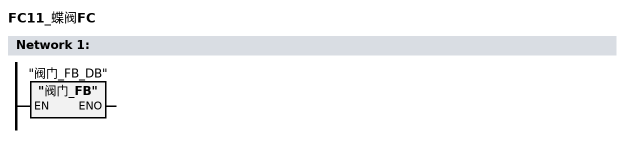
   RUNG wire#powerrail
      "阀门_FB_DB"()
   END_RUNG
   // the same network as SCL:
   "阀门_FB_DB"();   // "阀门_FB"
END_REGION
END_FUNCTION

FUNCTION "FC12_引水阀和排气阀FC" : Void   // FC12, LAD
{ S7_Optimized_Access := 'TRUE' }
VERSION : 0.1
BEGIN

REGION Network 1
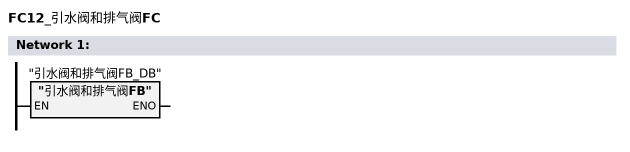
   RUNG wire#powerrail
      "引水阀和排气阀FB_DB"()
   END_RUNG
   // the same network as SCL:
   "引水阀和排气阀FB_DB"();   // "引水阀和排气阀FB"
END_REGION
END_FUNCTION

FUNCTION "FC13_电机_泵FC" : Void   // FC13, LAD
{ S7_Optimized_Access := 'TRUE' }
VERSION : 0.1
BEGIN

REGION Network 1
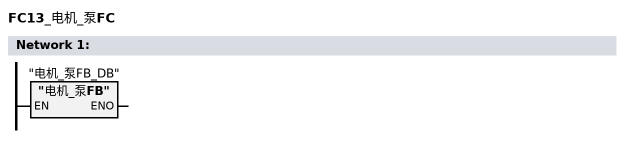
   RUNG wire#powerrail
      "电机_泵FB_DB"()
   END_RUNG
   // the same network as SCL:
   "电机_泵FB_DB"();   // "电机_泵FB"
END_REGION
END_FUNCTION

FUNCTION "FC14_DATA_ALARM" : Void   // FC14, LAD
{ S7_Optimized_Access := 'TRUE' }
VERSION : 0.1
BEGIN

REGION Network 1
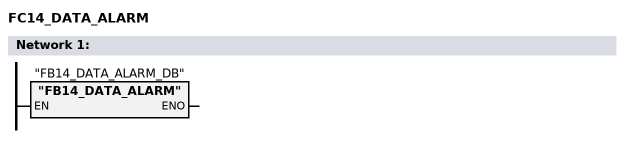
   RUNG wire#powerrail
      "FB14_DATA_ALARM_DB"()
   END_RUNG
   // the same network as SCL:
   "FB14_DATA_ALARM_DB"();   // "FB14_DATA_ALARM"
END_REGION
END_FUNCTION

FUNCTION "FC15_MOTOR_AUTO_ST" : Void   // FC15, LAD
{ S7_Optimized_Access := 'TRUE' }
VERSION : 0.1
BEGIN

REGION Network 1
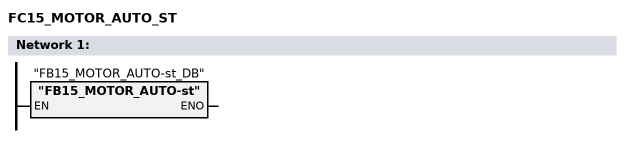
   RUNG wire#powerrail
      "FB15_MOTOR_AUTO-st_DB"()
   END_RUNG
   // the same network as SCL:
   "FB15_MOTOR_AUTO-st_DB"();   // "FB15_MOTOR_AUTO-st"
END_REGION
END_FUNCTION

FUNCTION "FC16" : Void   // FC16, LAD
{ S7_Optimized_Access := 'TRUE' }
VERSION : 0.1
   VAR_TEMP   // added for the SCL form of the ladder/FBD networks
      _w1 : Bool;
   END_VAR
BEGIN

REGION Network 1
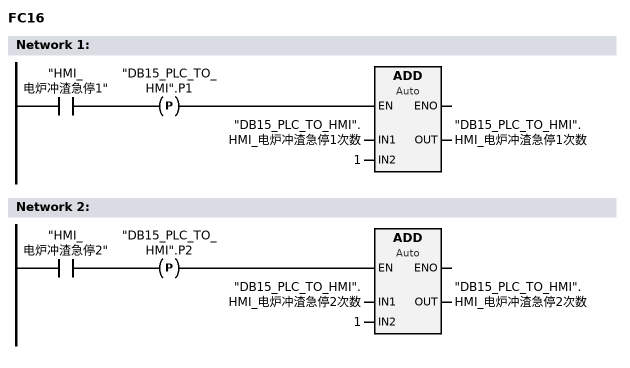
   RUNG wire#powerrail
      Contact( "HMI_电炉冲渣急停1" )
      P_Trig( "DB15_PLC_TO_HMI".P1 )
      Add(in1 := "DB15_PLC_TO_HMI".HMI_电炉冲渣急停1次数, in2 := 1, out => "DB15_PLC_TO_HMI".HMI_电炉冲渣急停1次数)
   END_RUNG
   // the same network as SCL:
   #_w1 := "HMI_电炉冲渣急停1" AND NOT "DB15_PLC_TO_HMI".P1;   // rising edge
   "DB15_PLC_TO_HMI".P1 := "HMI_电炉冲渣急停1";
   IF #_w1 THEN "DB15_PLC_TO_HMI".HMI_电炉冲渣急停1次数 := "DB15_PLC_TO_HMI".HMI_电炉冲渣急停1次数 + 1; END_IF;
END_REGION

REGION Network 2
   RUNG wire#powerrail
      Contact( "HMI_电炉冲渣急停2" )
      P_Trig( "DB15_PLC_TO_HMI".P2 )
      Add(in1 := "DB15_PLC_TO_HMI".HMI_电炉冲渣急停2次数, in2 := 1, out => "DB15_PLC_TO_HMI".HMI_电炉冲渣急停2次数)
   END_RUNG
   // the same network as SCL:
   #_w1 := "HMI_电炉冲渣急停2" AND NOT "DB15_PLC_TO_HMI".P2;   // rising edge
   "DB15_PLC_TO_HMI".P2 := "HMI_电炉冲渣急停2";
   IF #_w1 THEN "DB15_PLC_TO_HMI".HMI_电炉冲渣急停2次数 := "DB15_PLC_TO_HMI".HMI_电炉冲渣急停2次数 + 1; END_IF;
END_REGION
END_FUNCTION

ORGANIZATION_BLOCK "Main"   // OB1, LAD, ProgramCycle
TITLE = "Main Program Sweep (Cycle)"
{ S7_Optimized_Access := 'TRUE' }
VERSION : 0.1
   VAR_INPUT
      Initial_Call : Bool;   // Initial call of this OB
      Remanence : Bool;   // =True, if remanent data are available
   END_VAR
BEGIN

REGION Network 1
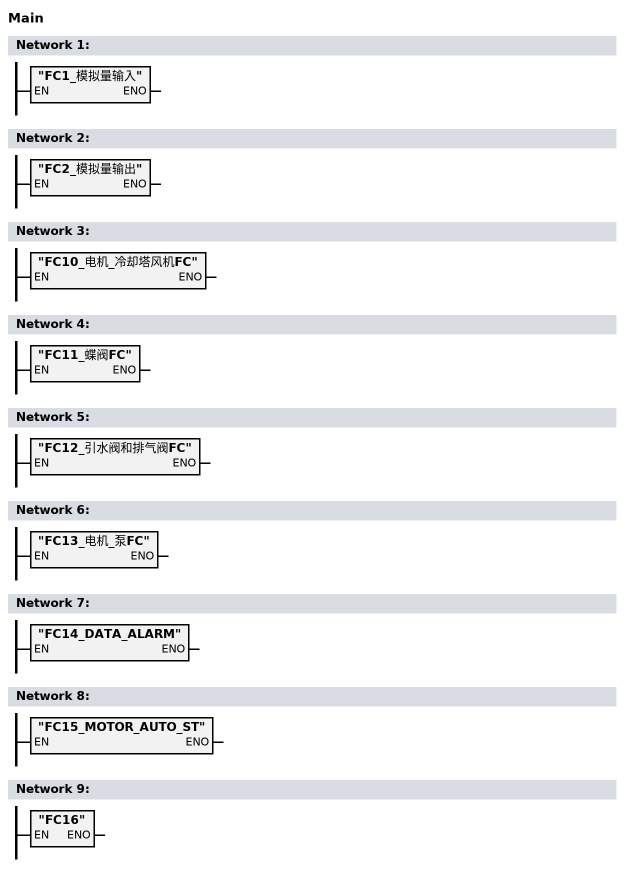
   RUNG wire#powerrail
      "FC1_模拟量输入"()
   END_RUNG
   // the same network as SCL:
   "FC1_模拟量输入"();
END_REGION

REGION Network 2
   RUNG wire#powerrail
      "FC2_模拟量输出"()
   END_RUNG
   // the same network as SCL:
   "FC2_模拟量输出"();
END_REGION

REGION Network 3
   RUNG wire#powerrail
      "FC10_电机_冷却塔风机FC"()
   END_RUNG
   // the same network as SCL:
   "FC10_电机_冷却塔风机FC"();
END_REGION

REGION Network 4
   RUNG wire#powerrail
      "FC11_蝶阀FC"()
   END_RUNG
   // the same network as SCL:
   "FC11_蝶阀FC"();
END_REGION

REGION Network 5
   RUNG wire#powerrail
      "FC12_引水阀和排气阀FC"()
   END_RUNG
   // the same network as SCL:
   "FC12_引水阀和排气阀FC"();
END_REGION

REGION Network 6
   RUNG wire#powerrail
      "FC13_电机_泵FC"()
   END_RUNG
   // the same network as SCL:
   "FC13_电机_泵FC"();
END_REGION

REGION Network 7
   RUNG wire#powerrail
      "FC14_DATA_ALARM"()
   END_RUNG
   // the same network as SCL:
   "FC14_DATA_ALARM"();
END_REGION

REGION Network 8
   RUNG wire#powerrail
      "FC15_MOTOR_AUTO_ST"()
   END_RUNG
   // the same network as SCL:
   "FC15_MOTOR_AUTO_ST"();
END_REGION

REGION Network 9
   RUNG wire#powerrail
      "FC16"()
   END_RUNG
   // the same network as SCL:
   "FC16"();
END_REGION
END_ORGANIZATION_BLOCK

ORGANIZATION_BLOCK "Cyclic interrupt"   // OB30, LAD, CyclicInterrupt
{ S7_Optimized_Access := 'TRUE' }
VERSION : 0.1
   VAR_INPUT
      Initial_Call : Bool;   // Initial call of this OB
      Event_Count : Int;   // Events discarded
   END_VAR
BEGIN
END_ORGANIZATION_BLOCK

// ===== PLC "2#SBF"  CPU 1511-1 PN =====

VAR_GLOBAL   // PLC tag table "默认变量表"
   "System_Byte" AT %MB1 : Byte;
   "FirstScan" AT %M1.0 : Bool;
   "DiagStatusUpdate" AT %M1.1 : Bool;
   "AlwaysTRUE" AT %M1.2 : Bool;
   "AlwaysFALSE" AT %M1.3 : Bool;
   "Clock_Byte" AT %MB0 : Byte;
   "Clock_10Hz" AT %M0.0 : Bool;
   "Clock_5Hz" AT %M0.1 : Bool;
   "Clock_2.5Hz" AT %M0.2 : Bool;
   "Clock_2Hz" AT %M0.3 : Bool;
   "Clock_1.25Hz" AT %M0.4 : Bool;
   "Clock_1Hz" AT %M0.5 : Bool;
   "Clock_0.625Hz" AT %M0.6 : Bool;
   "Clock_0.5Hz" AT %M0.7 : Bool;
   "1#冲渣泵本地/远程" AT %I0.0 : Bool;
   "1#冲渣泵备妥" AT %I0.1 : Bool;
   "1#冲渣泵运行" AT %I0.2 : Bool;
   "1#冲渣泵故障" AT %I0.3 : Bool;
   "2#冲渣泵本地/远程" AT %I0.4 : Bool;
   "2#冲渣泵备妥" AT %I0.5 : Bool;
   "2#冲渣泵运行" AT %I0.6 : Bool;
   "2#冲渣泵故障" AT %I0.7 : Bool;
   "3#冲渣泵本地/远程" AT %I1.0 : Bool;
   "3#冲渣泵备妥" AT %I1.1 : Bool;
   "3#冲渣泵运行" AT %I1.2 : Bool;
   "3#冲渣泵故障" AT %I1.3 : Bool;
   "4#冲渣泵本地/远程" AT %I1.4 : Bool;
   "4#冲渣泵备妥" AT %I1.5 : Bool;
   "4#冲渣泵运行" AT %I1.6 : Bool;
   "4#冲渣泵故障" AT %I1.7 : Bool;
   "5#冲渣泵本地/远程" AT %I2.0 : Bool;
   "5#冲渣泵备妥" AT %I2.1 : Bool;
   "5#冲渣泵运行" AT %I2.2 : Bool;
   "5#冲渣泵故障" AT %I2.3 : Bool;
   "6#冲渣泵本地/远程" AT %I2.4 : Bool;
   "6#冲渣泵备妥" AT %I2.5 : Bool;
   "6#冲渣泵运行" AT %I2.6 : Bool;
   "6#冲渣泵故障" AT %I2.7 : Bool;
   "7#冲渣泵本地/远程" AT %I3.0 : Bool;
   "7#冲渣泵备妥" AT %I3.1 : Bool;
   "7#冲渣泵运行" AT %I3.2 : Bool;
   "7#冲渣泵故障" AT %I3.3 : Bool;
   "8#冲渣泵本地/远程" AT %I3.4 : Bool;
   "8#冲渣泵备妥" AT %I3.5 : Bool;
   "8#冲渣泵运行" AT %I3.6 : Bool;
   "8#冲渣泵故障" AT %I3.7 : Bool;
   "1#热水泵本地/远程" AT %I4.0 : Bool;
   "1#热水泵备妥" AT %I4.1 : Bool;
   "1#热水泵运行" AT %I4.2 : Bool;
   "1#热水泵故障" AT %I4.3 : Bool;
   "2#热水泵本地/远程" AT %I4.4 : Bool;
   "2#热水泵备妥" AT %I4.5 : Bool;
   "2#热水泵运行" AT %I4.6 : Bool;
   "2#热水泵故障" AT %I4.7 : Bool;
   "3#热水泵本地/远程" AT %I5.0 : Bool;
   "3#热水泵备妥" AT %I5.1 : Bool;
   "3#热水泵运行" AT %I5.2 : Bool;
   "3#热水泵故障" AT %I5.3 : Bool;
   "4#热水泵本地/远程" AT %I5.4 : Bool;
   "4#热水泵备妥" AT %I5.5 : Bool;
   "4#热水泵运行" AT %I5.6 : Bool;
   "4#热水泵故障" AT %I5.7 : Bool;
   "5#热水泵本地/远程" AT %I6.0 : Bool;
   "5#热水泵备妥" AT %I6.1 : Bool;
   "5#热水泵运行" AT %I6.2 : Bool;
   "5#热水泵故障" AT %I6.3 : Bool;
   "6#热水泵本地/远程" AT %I6.4 : Bool;
   "6#热水泵备妥" AT %I6.5 : Bool;
   "6#热水泵运行" AT %I6.6 : Bool;
   "6#热水泵故障" AT %I6.7 : Bool;
   "7#热水泵本地/远程" AT %I7.0 : Bool;
   "7#热水泵备妥" AT %I7.1 : Bool;
   "7#热水泵运行" AT %I7.2 : Bool;
   "7#热水泵故障" AT %I7.3 : Bool;
   "8#热水泵本地/远程" AT %I7.4 : Bool;
   "8#热水泵备妥" AT %I7.5 : Bool;
   "8#热水泵运行" AT %I7.6 : Bool;
   "8#热水泵故障" AT %I7.7 : Bool;
   "1#浊环水上塔风机本地/远程" AT %I8.0 : Bool;
   "1#上塔风机备妥" AT %I8.1 : Bool;
   "1#上塔风机运行" AT %I8.2 : Bool;
   "1#上塔风机故障" AT %I8.3 : Bool;
   "2#浊环水上塔风机本地/远程" AT %I8.4 : Bool;
   "2#上塔风机备妥" AT %I8.5 : Bool;
   "2#上塔风机运行" AT %I8.6 : Bool;
   "2#上塔风机故障" AT %I8.7 : Bool;
   "3#浊环水上塔风机本地/远程" AT %I9.0 : Bool;
   "3#上塔风机备妥" AT %I9.1 : Bool;
   "3#上塔风机运行" AT %I9.2 : Bool;
   "3#上塔风机故障" AT %I9.3 : Bool;
   "4#浊环水上塔风机本地/远程" AT %I9.4 : Bool;
   "4#上塔风机备妥" AT %I9.5 : Bool;
   "4#上塔风机运行" AT %I9.6 : Bool;
   "4#上塔风机故障" AT %I9.7 : Bool;
   "5#浊环水上塔风机本地/远程" AT %I10.0 : Bool;
   "5#上塔风机备妥" AT %I10.1 : Bool;
   "5#上塔风机运行" AT %I10.2 : Bool;
   "5#上塔风机故障" AT %I10.3 : Bool;
   "6#浊环水上塔风机本地/远程" AT %I10.4 : Bool;
   "6#上塔风机备妥" AT %I10.5 : Bool;
   "6#上塔风机运行" AT %I10.6 : Bool;
   "6#上塔风机故障" AT %I10.7 : Bool;
   "1#炉体循环水泵本地/远程" AT %I11.0 : Bool;
   "1#炉体循环水泵备妥" AT %I11.1 : Bool;
   "1#炉体循环水泵运行" AT %I11.2 : Bool;
   "1#炉体循环水泵故障" AT %I11.3 : Bool;
   "2#炉体循环水泵本地/远程" AT %I11.4 : Bool;
   "2#炉体循环水泵备妥" AT %I11.5 : Bool;
   "2#炉体循环水泵运行" AT %I11.6 : Bool;
   "2#炉体循环水泵故障" AT %I11.7 : Bool;
   "3#炉体循环水泵本地/远程" AT %I12.0 : Bool;
   "3#炉体循环水泵备妥" AT %I12.1 : Bool;
   "3#炉体循环水泵运行" AT %I12.2 : Bool;
   "3#炉体循环水泵故障" AT %I12.3 : Bool;
   "1#电极冷却水泵本地/远程" AT %I12.4 : Bool;
   "1#电极冷却水泵备妥" AT %I12.5 : Bool;
   "1#电极冷却水泵运行" AT %I12.6 : Bool;
   "1#电极冷却水泵故障" AT %I12.7 : Bool;
   "2#电极冷却水泵本地/远程" AT %I13.0 : Bool;
   "2#电极冷却水泵备妥" AT %I13.1 : Bool;
   "2#电极冷却水泵运行" AT %I13.2 : Bool;
   "2#电极冷却水泵故障" AT %I13.3 : Bool;
   "3#电极冷却水泵本地/远程" AT %I13.4 : Bool;
   "3#电极冷却水泵备妥" AT %I13.5 : Bool;
   "3#电极冷却水泵运行" AT %I13.6 : Bool;
   "3#电极冷却水泵故障" AT %I13.7 : Bool;
   "4#电极冷却水泵本地/远程" AT %I14.0 : Bool;
   "4#电极冷却水泵备妥" AT %I14.1 : Bool;
   "4#电极冷却水泵运行" AT %I14.2 : Bool;
   "4#电极冷却水泵故障" AT %I14.3 : Bool;
   "1#净环热水泵本地/远程" AT %I14.4 : Bool;
   "1#净环热水泵备妥" AT %I14.5 : Bool;
   "1#净环热水泵运行" AT %I14.6 : Bool;
   "1#净环热水泵故障" AT %I14.7 : Bool;
   "2#净环热水泵本地/远程" AT %I15.0 : Bool;
   "2#净环热水泵备妥" AT %I15.1 : Bool;
   "2#净环热水泵运行" AT %I15.2 : Bool;
   "2#净环热水泵故障" AT %I15.3 : Bool;
   "3#净环热水泵本地/远程" AT %I15.4 : Bool;
   "3#净环热水泵备妥" AT %I15.5 : Bool;
   "3#净环热水泵运行" AT %I15.6 : Bool;
   "3#净环热水泵故障" AT %I15.7 : Bool;
   "4#净环热水泵本地/远程" AT %I16.0 : Bool;
   "4#净环热水泵备妥" AT %I16.1 : Bool;
   "4#净环热水泵运行" AT %I16.2 : Bool;
   "4#净环热水泵故障" AT %I16.3 : Bool;
   "5#净环热水泵本地/远程" AT %I16.4 : Bool;
   "5#净环热水泵备妥" AT %I16.5 : Bool;
   "5#净环热水泵运行" AT %I16.6 : Bool;
   "5#净环热水泵故障" AT %I16.7 : Bool;
   "1#柴油泵本地/远程" AT %I17.0 : Bool;
   "1#柴油泵备妥" AT %I17.1 : Bool;
   "1#柴油泵运行" AT %I17.2 : Bool;
   "1#柴油泵故障" AT %I17.3 : Bool;
   "2#柴油泵本地/远程" AT %I17.4 : Bool;
   "2#柴油泵备妥" AT %I17.5 : Bool;
   "2#柴油泵运行" AT %I17.6 : Bool;
   "2#柴油泵故障" AT %I17.7 : Bool;
   "1#净环上塔风机本地/远程" AT %I18.0 : Bool;
   "1#净环上塔风机备妥" AT %I18.1 : Bool;
   "1#净环上塔风机运行" AT %I18.2 : Bool;
   "1#净环上塔风机故障" AT %I18.3 : Bool;
   "2#净环上塔风机本地/远程" AT %I18.4 : Bool;
   "2#净环上塔风机备妥" AT %I18.5 : Bool;
   "2#净环上塔风机运行" AT %I18.6 : Bool;
   "2#净环上塔风机故障" AT %I18.7 : Bool;
   "3#净环上塔风机本地/远程" AT %I19.0 : Bool;
   "3#净环上塔风机备妥" AT %I19.1 : Bool;
   "3#净环上塔风机运行" AT %I19.2 : Bool;
   "3#净环上塔风机故障" AT %I19.3 : Bool;
   "窑冷却泵备妥" AT %I19.4 : Bool;
   "4#净环上塔风机备妥" AT %I19.5 : Bool;
   "4#净环上塔风机运行" AT %I19.6 : Bool;
   "4#净环上塔风机故障" AT %I19.7 : Bool;
   "1#冲渣泵空气监测" AT %I20.0 : Bool;
   "2#冲渣泵空气监测" AT %I20.1 : Bool;
   "3#冲渣泵空气监测" AT %I20.2 : Bool;
   "4#冲渣泵空气监测" AT %I20.3 : Bool;
   "5#冲渣泵空气监测" AT %I20.4 : Bool;
   "6#冲渣泵空气监测" AT %I20.5 : Bool;
   "7#冲渣泵空气监测" AT %I20.6 : Bool;
   "8#冲渣泵空气监测" AT %I20.7 : Bool;
   "1#浊环热水泵空气监测" AT %I21.0 : Bool;
   "2#浊环热水泵空气监测" AT %I21.1 : Bool;
   "3#浊环热水泵空气监测" AT %I21.2 : Bool;
   "4#浊环热水泵空气监测" AT %I21.3 : Bool;
   "5#浊环热水泵空气监测" AT %I21.4 : Bool;
   "6#浊环热水泵空气监测" AT %I21.5 : Bool;
   "7#浊环热水泵空气监测" AT %I21.6 : Bool;
   "8#浊环热水泵空气监测" AT %I21.7 : Bool;
   "1#炉体水泵空气监测" AT %I22.0 : Bool;
   "2#炉体水泵空气监测" AT %I22.1 : Bool;
   "3#炉体水泵空气监测" AT %I22.2 : Bool;
   "1#电极水泵空气监测" AT %I22.3 : Bool;
   "2#电极水泵空气监测" AT %I22.4 : Bool;
   "3#电极水泵空气监测" AT %I22.5 : Bool;
   "4#电极水泵空气监测" AT %I22.6 : Bool;
   "1#净环热水泵空气监测" AT %I22.7 : Bool;
   "2#净环热水泵空气监测" AT %I23.0 : Bool;
   "3#净环热水泵空气监测" AT %I23.1 : Bool;
   "4#净环热水泵空气监测" AT %I23.2 : Bool;
   "5#净环热水泵空气监测" AT %I23.3 : Bool;
   "1#柴油水泵空气监测" AT %I23.4 : Bool;
   "2#柴油水泵空气监测" AT %I23.5 : Bool;
   "1#冲渣泵驱动" AT %Q0.0 : Bool;
   "2#冲渣泵驱动" AT %Q0.1 : Bool;
   "3#冲渣泵驱动" AT %Q0.2 : Bool;
   "4#冲渣泵驱动" AT %Q0.3 : Bool;
   "5#冲渣泵驱动" AT %Q0.4 : Bool;
   "6#冲渣泵驱动" AT %Q0.5 : Bool;
   "7#冲渣泵驱动" AT %Q0.6 : Bool;
   "8#冲渣泵驱动" AT %Q0.7 : Bool;
   "1#浊环热水泵驱动" AT %Q1.0 : Bool;
   "2#浊环热水泵驱动" AT %Q1.1 : Bool;
   "3#浊环热水泵驱动" AT %Q1.2 : Bool;
   "4#浊环热水泵驱动" AT %Q1.3 : Bool;
   "5#浊环热水泵驱动" AT %Q1.4 : Bool;
   "6#浊环热水泵驱动" AT %Q1.5 : Bool;
   "7#浊环热水泵驱动" AT %Q1.6 : Bool;
   "8#浊环热水泵驱动" AT %Q1.7 : Bool;
   "1#浊环水上塔风机" AT %Q2.0 : Bool;
   "2#浊环水上塔风机" AT %Q2.1 : Bool;
   "3#浊环水上塔风机" AT %Q2.2 : Bool;
   "4#浊环水上塔风机" AT %Q2.3 : Bool;
   "5#浊环水上塔风机" AT %Q2.4 : Bool;
   "6#浊环水上塔风机" AT %Q2.5 : Bool;
   "1#炉体循环水泵驱动" AT %Q2.6 : Bool;
   "2#炉体循环水泵驱动" AT %Q2.7 : Bool;
   "3#炉体循环水泵驱动" AT %Q3.0 : Bool;
   "1#电极循环水泵驱动" AT %Q3.1 : Bool;
   "2#电极循环水泵驱动" AT %Q3.2 : Bool;
   "3#电极循环水泵驱动" AT %Q3.3 : Bool;
   "4#电极循环水泵驱动" AT %Q3.4 : Bool;
   "1#净环热水泵驱动" AT %Q3.5 : Bool;
   "2#净环热水泵驱动" AT %Q3.6 : Bool;
   "3#净环热水泵驱动" AT %Q3.7 : Bool;
   "4#净环热水泵驱动" AT %Q4.0 : Bool;
   "1#净环水上塔风机" AT %Q4.1 : Bool;
   "2#净环水上塔风机" AT %Q4.2 : Bool;
   "3#净环水上塔风机" AT %Q4.3 : Bool;
   "4#净环水上塔风机" AT %Q4.4 : Bool;
   "1#柴油泵驱动" AT %Q4.5 : Bool;
   "2#柴油泵驱动" AT %Q4.6 : Bool;
   "1#炉体循环水电动蝶阀备妥" AT %I24.0 : Bool;
   "1#炉体循环水电动蝶阀运行" AT %I24.1 : Bool;
   "1#炉体循环水电动蝶阀故障" AT %I24.2 : Bool;
   "1#炉体循环水电动蝶阀开到位" AT %I24.3 : Bool;
   "1#炉体循环水电动蝶阀关到位" AT %I24.4 : Bool;
   "2#炉体循环水电动蝶阀备妥" AT %I24.5 : Bool;
   "2#炉体循环水电动蝶阀运行" AT %I24.6 : Bool;
   "2#炉体循环水电动蝶阀故障" AT %I24.7 : Bool;
   "2#炉体循环水电动蝶阀开到位" AT %I25.0 : Bool;
   "2#炉体循环水电动蝶阀关到位" AT %I25.1 : Bool;
   "3#炉体循环水电动蝶阀备妥" AT %I25.2 : Bool;
   "3#炉体循环水电动蝶阀运行" AT %I25.3 : Bool;
   "3#炉体循环水电动蝶阀故障" AT %I25.4 : Bool;
   "3#炉体循环水电动蝶阀开到位" AT %I25.5 : Bool;
   "3#炉体循环水电动蝶阀关到位" AT %I25.6 : Bool;
   "1#电极冷却水电动蝶阀备妥" AT %I25.7 : Bool;
   "1#电极冷却水电动蝶阀运行" AT %I26.0 : Bool;
   "1#电极冷却水电动蝶阀故障" AT %I26.1 : Bool;
   "1#电极冷却水电动蝶阀开到位" AT %I26.2 : Bool;
   "1#电极冷却水电动蝶阀关到位" AT %I26.3 : Bool;
   "2#电极冷却水电动蝶阀备妥" AT %I26.4 : Bool;
   "2#电极冷却水电动蝶阀运行" AT %I26.5 : Bool;
   "2#电极冷却水电动蝶阀故障" AT %I26.6 : Bool;
   "2#电极冷却水电动蝶阀开到位" AT %I26.7 : Bool;
   "2#电极冷却水电动蝶阀关到位" AT %I27.0 : Bool;
   "3#电极冷却水电动蝶阀备妥" AT %I27.1 : Bool;
   "3#电极冷却水电动蝶阀运行" AT %I27.2 : Bool;
   "3#电极冷却水电动蝶阀故障" AT %I27.3 : Bool;
   "3#电极冷却水电动蝶阀开到位" AT %I27.4 : Bool;
   "3#电极冷却水电动蝶阀关到位" AT %I27.5 : Bool;
   "4#电极冷却水电动蝶阀备妥" AT %I27.6 : Bool;
   "4#电极冷却水电动蝶阀运行" AT %I27.7 : Bool;
   "4#电极冷却水电动蝶阀故障" AT %I28.0 : Bool;
   "4#电极冷却水电动蝶阀开到位" AT %I28.1 : Bool;
   "4#电极冷却水电动蝶阀关到位" AT %I28.2 : Bool;
   "1#净环热水电动蝶阀备妥" AT %I28.3 : Bool;
   "1#净环热水电动蝶阀运行" AT %I28.4 : Bool;
   "1#净环热水电动蝶阀故障" AT %I28.5 : Bool;
   "1#净环热水电动蝶阀开到位" AT %I28.6 : Bool;
   "1#净环热水电动蝶阀关到位" AT %I28.7 : Bool;
   "2#净环热水电动蝶阀备妥" AT %I29.0 : Bool;
   "2#净环热水电动蝶阀运行" AT %I29.1 : Bool;
   "2#净环热水电动蝶阀故障" AT %I29.2 : Bool;
   "2#净环热水电动蝶阀开到位" AT %I29.3 : Bool;
   "2#净环热水电动蝶阀关到位" AT %I29.4 : Bool;
   "3#净环热水电动蝶阀备妥" AT %I29.5 : Bool;
   "3#净环热水电动蝶阀运行" AT %I29.6 : Bool;
   "3#净环热水电动蝶阀故障" AT %I29.7 : Bool;
   "1#炉体循环水泵引水电磁阀" AT %Q8.0 : Bool;
   "3#净环热水电动蝶阀开到位" AT %I30.0 : Bool;
   "3#净环热水电动蝶阀关到位" AT %I30.1 : Bool;
   "4#净环热水电动蝶阀备妥" AT %I30.2 : Bool;
   "4#净环热水电动蝶阀运行" AT %I30.3 : Bool;
   "4#净环热水电动蝶阀故障" AT %I30.4 : Bool;
   "4#净环热水电动蝶阀开到位" AT %I30.5 : Bool;
   "4#净环热水电动蝶阀关到位" AT %I30.6 : Bool;
   "5#净环热水电动蝶阀备妥" AT %I30.7 : Bool;
   "5#净环热水电动蝶阀运行" AT %I31.0 : Bool;
   "5#净环热水电动蝶阀故障" AT %I31.1 : Bool;
   "5#净环热水电动蝶阀开到位" AT %I31.2 : Bool;
   "5#净环热水电动蝶阀关到位" AT %I31.3 : Bool;
   "1#柴油泵电动蝶阀备妥" AT %I31.4 : Bool;
   "1#柴油泵电动蝶阀运行" AT %I31.5 : Bool;
   "1#柴油泵电动蝶阀故障" AT %I31.6 : Bool;
   "1#柴油泵电动蝶阀开到位" AT %I31.7 : Bool;
   "1#柴油泵电动蝶阀关到位" AT %I32.0 : Bool;
   "2#柴油泵电动蝶阀备妥" AT %I32.1 : Bool;
   "2#柴油泵电动蝶阀运行" AT %I32.2 : Bool;
   "2#柴油泵电动蝶阀故障" AT %I32.3 : Bool;
   "2#柴油泵电动蝶阀开到位" AT %I32.4 : Bool;
   "2#柴油泵电动蝶阀关到位" AT %I32.5 : Bool;
   "1#炉体循环水泵电动阀开" AT %Q8.1 : Bool;
   "1#炉体循环水泵电动阀关" AT %Q8.2 : Bool;
   "1#炉体循环水泵排气电磁阀" AT %Q8.3 : Bool;
   "2#炉体循环水泵引水电磁阀" AT %Q8.4 : Bool;
   "2#炉体循环水泵电动阀开" AT %Q8.5 : Bool;
   "2#炉体循环水泵电动阀关" AT %Q8.6 : Bool;
   "2#炉体循环水泵排气电磁阀" AT %Q8.7 : Bool;
   "3#炉体循环水泵引水电磁阀" AT %Q9.0 : Bool;
   "3#炉体循环水泵电动阀开" AT %Q9.1 : Bool;
   "3#炉体循环水泵电动阀关" AT %Q9.2 : Bool;
   "3#炉体循环水泵排气电磁阀" AT %Q9.3 : Bool;
   "1#电极循环水泵引水电磁阀" AT %Q9.4 : Bool;
   "1#电极循环水泵电动阀开" AT %Q9.5 : Bool;
   "1#电极循环水泵电动阀关" AT %Q9.6 : Bool;
   "1#电极循环水泵排气电磁阀" AT %Q9.7 : Bool;
   "2#电极循环水泵引水电磁阀" AT %Q10.0 : Bool;
   "2#电极循环水泵电动阀开" AT %Q10.1 : Bool;
   "2#电极循环水泵电动阀关" AT %Q10.2 : Bool;
   "2#电极循环水泵排气电磁阀" AT %Q10.3 : Bool;
   "3#电极循环水泵引水电磁阀" AT %Q10.4 : Bool;
   "3#电极循环水泵电动阀开" AT %Q10.5 : Bool;
   "3#电极循环水泵电动阀关" AT %Q10.6 : Bool;
   "3#电极循环水泵排气电磁阀" AT %Q10.7 : Bool;
   "4#电极循环水泵引水电磁阀" AT %Q11.0 : Bool;
   "4#电极循环水泵电动阀开" AT %Q11.1 : Bool;
   "4#电极循环水泵电动阀关" AT %Q11.2 : Bool;
   "4#电极循环水泵排气电磁阀" AT %Q11.3 : Bool;
   "1#净环热水泵引水电磁阀" AT %Q11.4 : Bool;
   "1#净环热水泵电动阀开" AT %Q11.5 : Bool;
   "1#净环热水泵电动阀关" AT %Q11.6 : Bool;
   "1#净环热水泵排气电磁阀" AT %Q11.7 : Bool;
   "2#净环热水泵引水电磁阀" AT %Q12.0 : Bool;
   "2#净环热水泵电动阀开" AT %Q12.1 : Bool;
   "2#净环热水泵电动阀关" AT %Q12.2 : Bool;
   "2#净环热水泵排气电磁阀" AT %Q12.3 : Bool;
   "3#净环热水泵引水电磁阀" AT %Q12.4 : Bool;
   "3#净环热水泵电动阀开" AT %Q12.5 : Bool;
   "3#净环热水泵电动阀关" AT %Q12.6 : Bool;
   "3#净环热水泵排气电磁阀" AT %Q12.7 : Bool;
   "4#净环热水泵引水电磁阀" AT %Q13.0 : Bool;
   "4#净环热水泵电动阀开" AT %Q13.1 : Bool;
   "4#净环热水泵电动阀关" AT %Q13.2 : Bool;
   "4#净环热水泵排气电磁阀" AT %Q13.3 : Bool;
   "1#外围取水阀开" AT %Q13.4 : Bool;
   "1#外围取水阀关" AT %Q13.5 : Bool;
   "2#外围取水阀开" AT %Q13.6 : Bool;
   "2#外围取水阀关" AT %Q13.7 : Bool;
   "1#炉体水泵管道压力" AT %IW256 : Int;
   "2#炉体水泵管道压力" AT %IW258 : Int;
   "3#炉体水泵管道压力" AT %IW260 : Int;
   "1#电极水泵管道压力" AT %IW262 : Int;
   "2#电极水泵管道压力" AT %IW264 : Int;
   "3#电极水泵管道压力" AT %IW266 : Int;
   "4#电极水泵管道压力" AT %IW268 : Int;
   "1#柴油泵管道压力" AT %IW270 : Int;
   "2#柴油泵管道压力" AT %IW272 : Int;
   "1#炉体水阀门开度" AT %IW274 : Int;
   "2#炉体水阀门开度" AT %IW276 : Int;
   "3#炉体水阀门开度" AT %IW278 : Int;
   "1#电极水阀门开度" AT %IW280 : Int;
   "2#电极水阀门开度" AT %IW282 : Int;
   "3#电极水阀门开度" AT %IW284 : Int;
   "4#电极水阀门开度" AT %IW286 : Int;
   "2#柴油泵阀门开度" AT %IW288 : Int;
   "1#净环热水管道压力" AT %IW290 : Int;
   "2#净环热水管道压力" AT %IW292 : Int;
   "3#净环热水管道压力" AT %IW294 : Int;
   "4#净环热水管道压力" AT %IW296 : Int;
   "5#净环热水管道压力" AT %IW298 : Int;
   "6#净环热水管道压力" AT %IW300 : Int;
   "1#净环热水阀门开度" AT %IW302 : Int;
   "2#净环热水阀门开度" AT %IW304 : Int;
   "3#净环热水阀门开度" AT %IW306 : Int;
   "4#净环热水阀门开度" AT %IW308 : Int;
   "5#净环热水阀门开度" AT %IW310 : Int;
   "6#净环热水阀门开度" AT %IW312 : Int;
   "1#外围补水阀门开度" AT %IW314 : Int;
   "2#外围补水阀门开度" AT %IW316 : Int;
   "1#水池液位" AT %IW318 : Int;
   "2#水池液位" AT %IW320 : Int;
   "1#循环水泵阀门开度给定" AT %QW256 : Int;
   "2#循环水泵阀门开度给定" AT %QW258 : Int;
   "3#循环水泵阀门开度给定" AT %QW260 : Int;
   "1#电极冷却泵阀门开度给定" AT %QW262 : Int;
   "2#电极冷却泵阀门开度给定" AT %QW264 : Int;
   "3#电极冷却泵阀门开度给定" AT %QW266 : Int;
   "4#电极冷却泵阀门开度给定" AT %QW268 : Int;
   "1#柴油泵阀门开度给定" AT %QW270 : Int;
   "2#柴油泵阀门开度给定" AT %QW272 : Int;
   "1#净环热水泵阀门开度给定" AT %QW274 : Int;
   "2#净环热水泵阀门开度给定" AT %QW276 : Int;
   "3#净环热水泵阀门开度给定" AT %QW278 : Int;
   "4#净环热水泵阀门开度给定" AT %QW280 : Int;
   "5#净环热水泵阀门开度给定" AT %QW282 : Int;
   "6#净环热水泵阀门开度给定" AT %QW284 : Int;
   "1#外围补水阀门开度给定" AT %QW286 : Int;
   "2#外围补水阀门开度给定" AT %QW288 : Int;
   "1#热水电动蝶阀备妥" AT %I36.0 : Bool;
   "1#热水电动蝶阀运行" AT %I36.1 : Bool;
   "1#热水电动蝶阀故障" AT %I36.2 : Bool;
   "1#热水电动蝶阀开到位" AT %I36.3 : Bool;
   "1#热水电动蝶阀关到位" AT %I36.4 : Bool;
   "2#热水电动蝶阀备妥" AT %I36.5 : Bool;
   "2#热水电动蝶阀运行" AT %I36.6 : Bool;
   "2#热水电动蝶阀故障" AT %I36.7 : Bool;
   "2#热水电动蝶阀开到位" AT %I37.0 : Bool;
   "2#热水电动蝶阀关到位" AT %I37.1 : Bool;
   "3#热水电动蝶阀备妥" AT %I37.2 : Bool;
   "3#热水电动蝶阀运行" AT %I37.3 : Bool;
   "3#热水电动蝶阀故障" AT %I37.4 : Bool;
   "3#热水电动蝶阀开到位" AT %I37.5 : Bool;
   "3#热水电动蝶阀关到位" AT %I37.6 : Bool;
   "4#热水电动蝶阀备妥" AT %I37.7 : Bool;
   "4#热水电动蝶阀运行" AT %I38.0 : Bool;
   "4#热水电动蝶阀故障" AT %I38.1 : Bool;
   "4#热水电动蝶阀开到位" AT %I38.2 : Bool;
   "4#热水电动蝶阀关到位" AT %I38.3 : Bool;
   "5#热水电动蝶阀备妥" AT %I38.4 : Bool;
   "5#热水电动蝶阀运行" AT %I38.5 : Bool;
   "5#热水电动蝶阀故障" AT %I38.6 : Bool;
   "5#热水电动蝶阀开到位" AT %I38.7 : Bool;
   "5#热水电动蝶阀关到位" AT %I39.0 : Bool;
   "6#热水电动蝶阀备妥" AT %I39.1 : Bool;
   "6#热水电动蝶阀运行" AT %I39.2 : Bool;
   "6#热水电动蝶阀故障" AT %I39.3 : Bool;
   "6#热水电动蝶阀开到位" AT %I39.4 : Bool;
   "6#热水电动蝶阀关到位" AT %I39.5 : Bool;
   "7#热水电动蝶阀备妥" AT %I39.6 : Bool;
   "7#热水电动蝶阀运行" AT %I39.7 : Bool;
   "7#热水电动蝶阀故障" AT %I40.0 : Bool;
   "7#热水电动蝶阀开到位" AT %I40.1 : Bool;
   "7#热水电动蝶阀关到位" AT %I40.2 : Bool;
   "8#热水电动蝶阀备妥" AT %I40.3 : Bool;
   "8#热水电动蝶阀运行" AT %I40.4 : Bool;
   "8#热水电动蝶阀故障" AT %I40.5 : Bool;
   "8#热水电动蝶阀开到位" AT %I40.6 : Bool;
   "8#热水电动蝶阀关到位" AT %I40.7 : Bool;
   "1#浊环热水泵引水电磁阀" AT %Q16.0 : Bool;
   "1#浊环热水泵电动阀开" AT %Q16.1 : Bool;
   "1#浊环热水泵电动阀关" AT %Q16.2 : Bool;
   "1#浊环热水泵排气电磁阀" AT %Q16.3 : Bool;
   "2#浊环热水泵引水电磁阀" AT %Q16.4 : Bool;
   "2#浊环热水泵电动阀开" AT %Q16.5 : Bool;
   "2#浊环热水泵电动阀关" AT %Q16.6 : Bool;
   "2#浊环热水泵排气电磁阀" AT %Q16.7 : Bool;
   "3#浊环热水泵引水电磁阀" AT %Q17.0 : Bool;
   "3#浊环热水泵电动阀开" AT %Q17.1 : Bool;
   "3#浊环热水泵电动阀关" AT %Q17.2 : Bool;
   "3#浊环热水泵排气电磁阀" AT %Q17.3 : Bool;
   "4#浊环热水泵引水电磁阀" AT %Q17.4 : Bool;
   "4#浊环热水泵电动阀开" AT %Q17.5 : Bool;
   "4#浊环热水泵电动阀关" AT %Q17.6 : Bool;
   "4#浊环热水泵排气电磁阀" AT %Q17.7 : Bool;
   "5#浊环热水泵引水电磁阀" AT %Q18.0 : Bool;
   "5#浊环热水泵电动阀开" AT %Q18.1 : Bool;
   "5#浊环热水泵电动阀关" AT %Q18.2 : Bool;
   "5#浊环热水泵排气电磁阀" AT %Q18.3 : Bool;
   "6#浊环热水泵引水电磁阀" AT %Q18.4 : Bool;
   "6#浊环热水泵电动阀开" AT %Q18.5 : Bool;
   "6#浊环热水泵电动阀关" AT %Q18.6 : Bool;
   "6#浊环热水泵排气电磁阀" AT %Q18.7 : Bool;
   "7#浊环热水泵引水电磁阀" AT %Q19.0 : Bool;
   "7#浊环热水泵电动阀开" AT %Q19.1 : Bool;
   "7#浊环热水泵电动阀关" AT %Q19.2 : Bool;
   "7#浊环热水泵排气电磁阀" AT %Q19.3 : Bool;
   "8#浊环热水泵引水电磁阀" AT %Q19.4 : Bool;
   "8#浊环热水泵电动阀开" AT %Q19.5 : Bool;
   "8#浊环热水泵电动阀关" AT %Q19.6 : Bool;
   "8#浊环热水泵排气电磁阀" AT %Q19.7 : Bool;
   "1#冲渣热水泵管道压力" AT %IW336 : Int;
   "2#冲渣热水泵管道压力" AT %IW338 : Int;
   "3#冲渣热水泵管道压力" AT %IW340 : Int;
   "4#冲渣热水泵管道压力" AT %IW342 : Int;
   "5#冲渣热水泵管道压力" AT %IW344 : Int;
   "6#冲渣热水泵管道压力" AT %IW346 : Int;
   "7#冲渣热水泵管道压力" AT %IW348 : Int;
   "8#冲渣热水泵管道压力" AT %IW350 : Int;
   "1#冲渣热水阀门开度" AT %IW352 : Int;
   "2#冲渣热水阀门开度" AT %IW354 : Int;
   "3#冲渣热水阀门开度" AT %IW356 : Int;
   "4#冲渣热水阀门开度" AT %IW358 : Int;
   "5#冲渣热水阀门开度" AT %IW360 : Int;
   "6#冲渣热水阀门开度" AT %IW362 : Int;
   "7#冲渣热水阀门开度" AT %IW364 : Int;
   "8#冲渣热水阀门开度" AT %IW366 : Int;
   "1#冲渣热水泵阀门开度给定" AT %QW304 : Int;
   "2#冲渣热水泵阀门开度给定" AT %QW306 : Int;
   "3#冲渣热水泵阀门开度给定" AT %QW308 : Int;
   "4#冲渣热水泵阀门开度给定" AT %QW310 : Int;
   "5#冲渣热水泵阀门开度给定" AT %QW312 : Int;
   "6#冲渣热水泵阀门开度给定" AT %QW314 : Int;
   "7#冲渣热水泵阀门开度给定" AT %QW316 : Int;
   "8#冲渣热水泵阀门开度给定" AT %QW318 : Int;
   "1#冲渣电动蝶阀备妥" AT %I44.0 : Bool;
   "1#冲渣电动蝶阀运行" AT %I44.1 : Bool;
   "1#冲渣电动蝶阀故障" AT %I44.2 : Bool;
   "1#冲渣电动蝶阀开到位" AT %I44.3 : Bool;
   "1#冲渣电动蝶阀关到位" AT %I44.4 : Bool;
   "2#冲渣电动蝶阀备妥" AT %I44.5 : Bool;
   "2#冲渣电动蝶阀运行" AT %I44.6 : Bool;
   "2#冲渣电动蝶阀故障" AT %I44.7 : Bool;
   "2#冲渣电动蝶阀开到位" AT %I45.0 : Bool;
   "2#冲渣电动蝶阀关到位" AT %I45.1 : Bool;
   "3#冲渣电动蝶阀备妥" AT %I45.2 : Bool;
   "3#冲渣电动蝶阀运行" AT %I45.3 : Bool;
   "3#冲渣电动蝶阀故障" AT %I45.4 : Bool;
   "3#冲渣电动蝶阀开到位" AT %I45.5 : Bool;
   "3#冲渣电动蝶阀关到位" AT %I45.6 : Bool;
   "4#冲渣电动蝶阀备妥" AT %I45.7 : Bool;
   "4#冲渣电动蝶阀运行" AT %I46.0 : Bool;
   "4#冲渣电动蝶阀故障" AT %I46.1 : Bool;
   "4#冲渣电动蝶阀开到位" AT %I46.2 : Bool;
   "4#冲渣电动蝶阀关到位" AT %I46.3 : Bool;
   "5#冲渣电动蝶阀备妥" AT %I46.4 : Bool;
   "5#冲渣电动蝶阀运行" AT %I46.5 : Bool;
   "5#冲渣电动蝶阀故障" AT %I46.6 : Bool;
   "5#冲渣电动蝶阀开到位" AT %I46.7 : Bool;
   "5#冲渣电动蝶阀关到位" AT %I47.0 : Bool;
   "6#冲渣电动蝶阀备妥" AT %I47.1 : Bool;
   "6#冲渣电动蝶阀运行" AT %I47.2 : Bool;
   "6#冲渣电动蝶阀故障" AT %I47.3 : Bool;
   "6#冲渣电动蝶阀开到位" AT %I47.4 : Bool;
   "6#冲渣电动蝶阀关到位" AT %I47.5 : Bool;
   "7#冲渣电动蝶阀备妥" AT %I47.6 : Bool;
   "7#冲渣电动蝶阀运行" AT %I47.7 : Bool;
   "7#冲渣电动蝶阀故障" AT %I48.0 : Bool;
   "7#冲渣电动蝶阀开到位" AT %I48.1 : Bool;
   "7#冲渣电动蝶阀关到位" AT %I48.2 : Bool;
   "8#冲渣电动蝶阀备妥" AT %I48.3 : Bool;
   "8#冲渣电动蝶阀运行" AT %I48.4 : Bool;
   "8#冲渣电动蝶阀故障" AT %I48.5 : Bool;
   "8#冲渣电动蝶阀开到位" AT %I48.6 : Bool;
   "8#冲渣电动蝶阀关到位" AT %I48.7 : Bool;
   "1#冲渣泵引水电磁阀" AT %Q20.0 : Bool;
   "1#冲渣泵电动阀开" AT %Q20.1 : Bool;
   "1#冲渣泵电动阀关" AT %Q20.2 : Bool;
   "1#冲渣泵排气电磁阀" AT %Q20.3 : Bool;
   "2#冲渣泵引水电磁阀" AT %Q20.4 : Bool;
   "2#冲渣泵电动阀开" AT %Q20.5 : Bool;
   "2#冲渣泵电动阀关" AT %Q20.6 : Bool;
   "2#冲渣泵排气电磁阀" AT %Q20.7 : Bool;
   "3#冲渣泵引水电磁阀" AT %Q21.0 : Bool;
   "3#冲渣泵电动阀开" AT %Q21.1 : Bool;
   "3#冲渣泵电动阀关" AT %Q21.2 : Bool;
   "3#冲渣泵排气电磁阀" AT %Q21.3 : Bool;
   "4#冲渣泵引水电磁阀" AT %Q21.4 : Bool;
   "4#冲渣泵电动阀开" AT %Q21.5 : Bool;
   "4#冲渣泵电动阀关" AT %Q21.6 : Bool;
   "4#冲渣泵排气电磁阀" AT %Q21.7 : Bool;
   "5#冲渣泵引水电磁阀" AT %Q22.0 : Bool;
   "5#冲渣泵电动阀开" AT %Q22.1 : Bool;
   "5#冲渣泵电动阀关" AT %Q22.2 : Bool;
   "5#冲渣泵排气电磁阀" AT %Q22.3 : Bool;
   "6#冲渣泵引水电磁阀" AT %Q22.4 : Bool;
   "6#冲渣泵电动阀开" AT %Q22.5 : Bool;
   "6#冲渣泵电动阀关" AT %Q22.6 : Bool;
   "6#冲渣泵排气电磁阀" AT %Q22.7 : Bool;
   "7#冲渣泵引水电磁阀" AT %Q23.0 : Bool;
   "7#冲渣泵电动阀开" AT %Q23.1 : Bool;
   "7#冲渣泵电动阀关" AT %Q23.2 : Bool;
   "7#冲渣泵排气电磁阀" AT %Q23.3 : Bool;
   "8#冲渣泵引水电磁阀" AT %Q23.4 : Bool;
   "8#冲渣泵电动阀开" AT %Q23.5 : Bool;
   "8#冲渣泵电动阀关" AT %Q23.6 : Bool;
   "8#冲渣泵排气电磁阀" AT %Q23.7 : Bool;
   "1#冲渣泵管道压力" AT %IW368 : Int;
   "2#冲渣泵管道压力" AT %IW370 : Int;
   "3#冲渣泵管道压力" AT %IW372 : Int;
   "4#冲渣泵管道压力" AT %IW374 : Int;
   "5#冲渣泵管道压力" AT %IW376 : Int;
   "6#冲渣泵管道压力" AT %IW378 : Int;
   "7#冲渣泵管道压力" AT %IW380 : Int;
   "8#冲渣泵管道压力" AT %IW382 : Int;
   "1#冲渣阀门开度" AT %IW384 : Int;
   "2#冲渣阀门开度" AT %IW386 : Int;
   "3#冲渣阀门开度" AT %IW388 : Int;
   "4#冲渣阀门开度" AT %IW390 : Int;
   "5#冲渣阀门开度" AT %IW392 : Int;
   "6#冲渣阀门开度" AT %IW394 : Int;
   "7#冲渣阀门开度" AT %IW396 : Int;
   "8#冲渣阀门开度" AT %IW398 : Int;
   "1#冲渣泵阀门开度给定" AT %QW320 : Int;
   "2#冲渣泵阀门开度给定" AT %QW322 : Int;
   "3#冲渣泵阀门开度给定" AT %QW324 : Int;
   "4#冲渣泵阀门开度给定" AT %QW326 : Int;
   "5#冲渣泵阀门开度给定" AT %QW328 : Int;
   "6#冲渣泵阀门开度给定" AT %QW330 : Int;
   "7#冲渣泵阀门开度给定" AT %QW332 : Int;
   "8#冲渣泵阀门开度给定" AT %QW334 : Int;
   "窑冷却泵运行" AT %I23.6 : Bool;
   "窑冷却泵故障" AT %I23.7 : Bool;
   "窑冷却泵驱动" AT %Q4.7 : Bool;
   "Q5_0" AT %Q5.0 : Bool;
   "Q5_1" AT %Q5.1 : Bool;
   "Q5_2" AT %Q5.2 : Bool;
   "Q5_3" AT %Q5.3 : Bool;
   "Q5_4" AT %Q5.4 : Bool;
   "Q5_5" AT %Q5.5 : Bool;
   "Q5_6" AT %Q5.6 : Bool;
   "Q5_7" AT %Q5.7 : Bool;
   "Q6_0" AT %Q6.0 : Bool;
   "Q6_1" AT %Q6.1 : Bool;
   "Q6_2" AT %Q6.2 : Bool;
   "Q6_3" AT %Q6.3 : Bool;
   "Q6_4" AT %Q6.4 : Bool;
   "Q6_5" AT %Q6.5 : Bool;
   "Q6_6" AT %Q6.6 : Bool;
   "Q6_7" AT %Q6.7 : Bool;
   "Q7_0" AT %Q7.0 : Bool;
   "Q7_1" AT %Q7.1 : Bool;
   "Q7_2" AT %Q7.2 : Bool;
   "Q7_3" AT %Q7.3 : Bool;
   "Q7_4" AT %Q7.4 : Bool;
   "Q7_5" AT %Q7.5 : Bool;
   "Q7_6" AT %Q7.6 : Bool;
   "Q7_7" AT %Q7.7 : Bool;
   "I32_6" AT %I32.6 : Bool;
   "I32_7" AT %I32.7 : Bool;
   "I33_0" AT %I33.0 : Bool;
   "I33_1" AT %I33.1 : Bool;
   "I33_2" AT %I33.2 : Bool;
   "I33_3" AT %I33.3 : Bool;
   "I33_4" AT %I33.4 : Bool;
   "I33_5" AT %I33.5 : Bool;
   "I33_6" AT %I33.6 : Bool;
   "I33_7" AT %I33.7 : Bool;
   "I34_0" AT %I34.0 : Bool;
   "I34_1" AT %I34.1 : Bool;
   "I34_2" AT %I34.2 : Bool;
   "I34_3" AT %I34.3 : Bool;
   "I34_4" AT %I34.4 : Bool;
   "I34_5" AT %I34.5 : Bool;
   "I34_6" AT %I34.6 : Bool;
   "I34_7" AT %I34.7 : Bool;
   "I35_0" AT %I35.0 : Bool;
   "I35_1" AT %I35.1 : Bool;
   "I35_2" AT %I35.2 : Bool;
   "I35_3" AT %I35.3 : Bool;
   "I35_4" AT %I35.4 : Bool;
   "I35_5" AT %I35.5 : Bool;
   "I35_6" AT %I35.6 : Bool;
   "I35_7" AT %I35.7 : Bool;
   "Q14_0" AT %Q14.0 : Bool;
   "Q14_1" AT %Q14.1 : Bool;
   "Q14_2" AT %Q14.2 : Bool;
   "Q14_3" AT %Q14.3 : Bool;
   "Q14_4" AT %Q14.4 : Bool;
   "Q14_5" AT %Q14.5 : Bool;
   "Q14_6" AT %Q14.6 : Bool;
   "Q14_7" AT %Q14.7 : Bool;
   "Q15_0" AT %Q15.0 : Bool;
   "Q15_1" AT %Q15.1 : Bool;
   "Q15_2" AT %Q15.2 : Bool;
   "Q15_3" AT %Q15.3 : Bool;
   "Q15_4" AT %Q15.4 : Bool;
   "Q15_5" AT %Q15.5 : Bool;
   "Q15_6" AT %Q15.6 : Bool;
   "Q15_7" AT %Q15.7 : Bool;
   "PIW322" AT %IW322 : Int;
   "PIW324" AT %IW324 : Int;
   "PIW326" AT %IW326 : Int;
   "PIW328" AT %IW328 : Int;
   "PIW330" AT %IW330 : Int;
   "PIW332" AT %IW332 : Int;
   "PIW334" AT %IW334 : Int;
   "PQW290" AT %QW290 : Int;
   "PQW292" AT %QW292 : Int;
   "PQW294" AT %QW294 : Int;
   "PQW296" AT %QW296 : Int;
   "PQW298" AT %QW298 : Int;
   "PQW330" AT %QW300 : Int;
   "PQW332" AT %QW302 : Int;
   "I41_0" AT %I41.0 : Bool;
   "I41_1" AT %I41.1 : Bool;
   "I41_2" AT %I41.2 : Bool;
   "I41_3" AT %I41.3 : Bool;
   "I41_4" AT %I41.4 : Bool;
   "I41_5" AT %I41.5 : Bool;
   "I41_6" AT %I41.6 : Bool;
   "I41_7" AT %I41.7 : Bool;
   "I42_0" AT %I42.0 : Bool;
   "I42_1" AT %I42.1 : Bool;
   "I42_2" AT %I42.2 : Bool;
   "I42_3" AT %I42.3 : Bool;
   "I42_4" AT %I42.4 : Bool;
   "I42_5" AT %I42.5 : Bool;
   "I42_6" AT %I42.6 : Bool;
   "I42_7" AT %I42.7 : Bool;
   "I43_0" AT %I43.0 : Bool;
   "I43_1" AT %I43.1 : Bool;
   "I43_2" AT %I43.2 : Bool;
   "I43_3" AT %I43.3 : Bool;
   "I43_4" AT %I43.4 : Bool;
   "I43_5" AT %I43.5 : Bool;
   "I43_6" AT %I43.6 : Bool;
   "I43_7" AT %I43.7 : Bool;
   "I49_0" AT %I49.0 : Bool;
   "I49_1" AT %I49.1 : Bool;
   "I49_2" AT %I49.2 : Bool;
   "I49_3" AT %I49.3 : Bool;
   "I49_4" AT %I49.4 : Bool;
   "I49_5" AT %I49.5 : Bool;
   "I49_6" AT %I49.6 : Bool;
   "I49_7" AT %I49.7 : Bool;
   "I50_0" AT %I50.0 : Bool;
   "I50_1" AT %I50.1 : Bool;
   "I50_2" AT %I50.2 : Bool;
   "I50_3" AT %I50.3 : Bool;
   "I50_4" AT %I50.4 : Bool;
   "I50_5" AT %I50.5 : Bool;
   "I50_6" AT %I50.6 : Bool;
   "I50_7" AT %I50.7 : Bool;
   "I51_0" AT %I51.0 : Bool;
   "I51_1" AT %I51.1 : Bool;
   "I51_2" AT %I51.2 : Bool;
   "I51_3" AT %I51.3 : Bool;
   "I51_4" AT %I51.4 : Bool;
   "I51_5" AT %I51.5 : Bool;
   "I51_6" AT %I51.6 : Bool;
   "I51_7" AT %I51.7 : Bool;
END_VAR

// ===== PLC "2#LM"  CPU 1511-1 PN =====
